
screen "eProC - Seguimiento Datos" 1280x768, template "Template"
   TextField "Campo de texto_9" at 88,77 size 35x18; Text 'Araña'
   TextField "Campo de texto_10" at 265,77 size 32x18; Text 'Rolos'
   TextField "Campo de texto_11" at 439,77 size 54x18; Text 'Perfilador'
   TextField "Campo de texto_12" at 788,77 size 31x18; Text 'Pinza'
   TextField "Campo de texto_13" at 967,77 size 57x18; Text 'Plegadora'
   TextField "Campo de texto_16" at 88,130 size 12x18; Text 'A'
   IOField "Champ E/S_8" at 109,127 size 54x25; FormatPattern 9999999
      Appearance <- "Araña\Araña.PresenciaPieza"
      ProcessValue <- "Araña\Araña.A"
   IOField "Champ E/S_9" at 109,147 size 54x25; FormatPattern 9999999
      Appearance <- "Araña\Araña.PresenciaPieza"
      ProcessValue <- "Araña\Araña.B"
   IOField "Champ E/S_10" at 109,168 size 54x24; FormatPattern 9999999
      Appearance <- "Araña\Araña.PresenciaPieza"
      ProcessValue <- "Araña\Araña.C"
   IOField "Champ E/S_11" at 109,187 size 54x25; FormatPattern 9999999
      Appearance <- "Araña\Araña.PresenciaPieza"
      ProcessValue <- "Araña\Araña.D"
   TextField "Campo de texto_17" at 89,148 size 11x18; Text 'B'
   TextField "Campo de texto_18" at 89,168 size 11x18; Text 'C'
   TextField "Campo de texto_19" at 89,188 size 12x18; Text 'D'
   TextField "Campo de texto_20" at 265,131 size 12x18; Text 'A'
   IOField "Champ E/S_12" at 284,127 size 54x25; FormatPattern 9999999
      Appearance <- "Rolos\Rolos.PresenciaPieza"
      ProcessValue <- "Rolos\Rolos.A"
   IOField "Champ E/S_13" at 284,147 size 54x25; FormatPattern 9999999
      Appearance <- "Rolos\Rolos.PresenciaPieza"
      ProcessValue <- "Rolos\Rolos.B"
   IOField "Champ E/S_14" at 284,168 size 54x24; FormatPattern 9999999
      Appearance <- "Rolos\Rolos.PresenciaPieza"
      ProcessValue <- "Rolos\Rolos.C"
   IOField "Champ E/S_15" at 284,187 size 54x25; FormatPattern 9999999
      Appearance <- "Rolos\Rolos.PresenciaPieza"
      ProcessValue <- "Rolos\Rolos.D"
   TextField "Campo de texto_21" at 265,149 size 11x18; Text 'B'
   TextField "Campo de texto_22" at 265,169 size 11x18; Text 'C'
   TextField "Campo de texto_23" at 265,189 size 12x18; Text 'D'
   TextField "Campo de texto_24" at 439,131 size 12x18; Text 'A'
   IOField "Champ E/S_16" at 462,127 size 53x25; FormatPattern 9999999
      Appearance <- "Perfiladores\Perfilador.PresenciaPieza"
      ProcessValue <- "Perfiladores\Perfilador.A"
   IOField "Champ E/S_17" at 462,147 size 53x25; FormatPattern 9999999
      Appearance <- "Perfiladores\Perfilador.PresenciaPieza"
      ProcessValue <- "Perfiladores\Perfilador.B"
   IOField "Champ E/S_18" at 462,168 size 53x24; FormatPattern 9999999
      Appearance <- "Perfiladores\Perfilador.PresenciaPieza"
      ProcessValue <- "Perfiladores\Perfilador.C"
   IOField "Champ E/S_19" at 462,187 size 53x25; FormatPattern 9999999
      Appearance <- "Perfiladores\Perfilador.PresenciaPieza"
      ProcessValue <- "Perfiladores\Perfilador.D"
   TextField "Campo de texto_25" at 441,149 size 11x18; Text 'B'
   TextField "Campo de texto_26" at 441,169 size 11x18; Text 'C'
   TextField "Campo de texto_27" at 441,189 size 12x18; Text 'D'
   TextField "Campo de texto_28" at 788,131 size 12x18; Text 'A'
   IOField "Champ E/S_20" at 813,127 size 53x25; FormatPattern 9999999
      Appearance <- "Pinza\Pinza.PresenciaPieza"
      ProcessValue <- "Pinza\Pinza.A"
   IOField "Champ E/S_21" at 813,147 size 53x25; FormatPattern 9999999
      Appearance <- "Pinza\Pinza.PresenciaPieza"
      ProcessValue <- "Pinza\Pinza.B"
   IOField "Champ E/S_22" at 813,168 size 53x24; FormatPattern 9999999
      Appearance <- "Pinza\Pinza.PresenciaPieza"
      ProcessValue <- "Pinza\Pinza.C"
   IOField "Champ E/S_23" at 813,187 size 53x25; FormatPattern 9999999
      Appearance <- "Pinza\Pinza.PresenciaPieza"
      ProcessValue <- "Pinza\Pinza.D"
   TextField "Campo de texto_29" at 788,149 size 11x18; Text 'B'
   TextField "Campo de texto_30" at 788,169 size 11x18; Text 'C'
   TextField "Campo de texto_31" at 788,189 size 12x18; Text 'D'
   TextField "Campo de texto_32" at 967,131 size 12x18; Text 'A'
   IOField "Champ E/S_24" at 988,127 size 53x25; FormatPattern 9999999
      Appearance <- "Plegadora\Plegadora.PresenciaPieza"
      ProcessValue <- "Plegadora\Plegadora.A"
   IOField "Champ E/S_25" at 988,147 size 53x25; FormatPattern 9999999
      Appearance <- "Plegadora\Plegadora.PresenciaPieza"
      ProcessValue <- "Plegadora\Plegadora.B"
   IOField "Champ E/S_26" at 988,168 size 53x24; FormatPattern 9999999
      Appearance <- "Plegadora\Plegadora.PresenciaPieza"
      ProcessValue <- "Plegadora\Plegadora.C"
   IOField "Champ E/S_27" at 988,187 size 53x25; FormatPattern 9999999
      Appearance <- "Plegadora\Plegadora.PresenciaPieza"
      ProcessValue <- "Plegadora\Plegadora.D"
   TextField "Campo de texto_33" at 967,149 size 11x18; Text 'B'
   TextField "Campo de texto_34" at 967,169 size 11x18; Text 'C'
   TextField "Campo de texto_35" at 967,189 size 12x18; Text 'D'
   Button "Botón_8" at 437,38 size 80x36; TextOff 'Borrar'; PictureOff "Borrar Pulsador"
      on Click: ResetBit("Perfiladores\Perfilador.PresenciaPieza")
      Visibility <- "Perfiladores\Perfilador.PresenciaPieza"
   Button "Botón_9" at 263,38 size 80x36; TextOff 'Borrar'; PictureOff "Borrar Pulsador"
      on Click: ResetBit("Rolos\Rolos.PresenciaPieza")
      Visibility <- "Rolos\Rolos.PresenciaPieza"
   Button "Botón_10" at 86,38 size 80x36; TextOff 'Borrar'; PictureOff "Borrar Pulsador"
      on Click: ResetBit("Araña\Araña.PresenciaPieza")
      Visibility <- "Araña\Araña.PresenciaPieza"
   TextField "Campo de texto_113" at 615,77 size 31x18; Text 'Cinta'
   TextField "Campo de texto_114" at 615,131 size 12x18; Text 'A'
   IOField "Champ E/S_106" at 638,127 size 53x25; FormatPattern 9999999
      Appearance <- "Cinta\Cinta.PresenciaPieza"
      ProcessValue <- "Cinta\Cinta.A"
   IOField "Champ E/S_107" at 638,147 size 53x25; FormatPattern 9999999
      Appearance <- "Cinta\Cinta.PresenciaPieza"
      ProcessValue <- "Cinta\Cinta.B"
   IOField "Champ E/S_108" at 638,168 size 53x24; FormatPattern 9999999
      Appearance <- "Cinta\Cinta.PresenciaPieza"
      ProcessValue <- "Cinta\Cinta.C"
   IOField "Champ E/S_109" at 638,187 size 53x25; FormatPattern 9999999
      Appearance <- "Cinta\Cinta.PresenciaPieza"
      ProcessValue <- "Cinta\Cinta.D"
   TextField "Campo de texto_115" at 615,149 size 11x18; Text 'B'
   TextField "Campo de texto_116" at 615,169 size 11x18; Text 'C'
   TextField "Campo de texto_117" at 615,189 size 12x18; Text 'D'
   Button "Botón_14" at 613,38 size 80x36; TextOff 'Borrar'; PictureOff "Borrar Pulsador"
      on Click: ResetBit("Cinta\Cinta.PresenciaPieza")
      Visibility <- "Cinta\Cinta.PresenciaPieza"
   Button "Botón_15" at 788,38 size 80x36; TextOff 'Borrar'; PictureOff "Borrar Pulsador"
      on Click: ResetBit("Pinza\Pinza.PresenciaPieza")
      Visibility <- "Pinza\Pinza.PresenciaPieza"
   Button "Botón_16" at 963,38 size 80x36; TextOff 'Borrar'; PictureOff "Borrar Pulsador"
      on Click: ResetBit("Plegadora\Plegadora.PresenciaPieza")
      Visibility <- "Plegadora\Plegadora.PresenciaPieza"
   GraphicView "Visor de gráficos_2" at 211,77 size 29x29; Picture "Gráfico_4"
   GraphicView "Visor de gráficos_1" at 384,77 size 29x29; Picture "Gráfico_4"
   GraphicView "Visor de gráficos_3" at 561,77 size 29x29; Picture "Gráfico_4"
   GraphicView "Visor de gráficos_4" at 734,77 size 29x29; Picture "Gráfico_4"
   GraphicView "Visor de gráficos_5" at 909,77 size 29x29; Picture "Gráfico_4"
   TextField "Campo de texto_1" at 72,425 size 54x29; Text 'Pinza'
   TextField "Campo de texto_2" at 229,507 size 54x18; Text 'Solicitada'
   TextField "Campo de texto_49" at 142,529 size 60x18; Text 'Recepción'
   IOField "Champ E/S_1" at 221,525 size 85x25; FormatPattern s9999999999
      ProcessValue <- "Pos_Recepcion"
      Appearance <- "Pinza\Pinza.PresenciaPieza"
   IOField "Champ E/S_2" at 221,545 size 85x25; FormatPattern s9999999999
      ProcessValue <- "Pos_E1H1"
      Appearance <- "Pinza\Pinza.PresenciaPieza"
   IOField "Champ E/S_3" at 221,566 size 85x24; FormatPattern s9999999999
      ProcessValue <- "Pos_E1H2"
      Appearance <- "Pinza\Pinza.PresenciaPieza"
   IOField "Champ E/S_4" at 221,585 size 85x25; FormatPattern s9999999999
      ProcessValue <- "Pos_E2H1"
      Appearance <- "Pinza\Pinza.PresenciaPieza"
   TextField "Campo de texto_50" at 142,547 size 33x18; Text 'E1H1'
   TextField "Campo de texto_51" at 142,567 size 33x18; Text 'E1H2'
   TextField "Campo de texto_52" at 142,587 size 33x18; Text 'E2H1'
   TextField "Campo de texto_53" at 313,507 size 57x18; Text 'Alcanzada'
   IOField "Champ E/S_5" at 305,525 size 85x25; FormatPattern s9999999999
      ProcessValue <- "Pos_Recepcion(3)"
      Appearance <- "Pinza\Pinza.PresenciaPieza"
   IOField "Champ E/S_6" at 305,545 size 85x25; FormatPattern s9999999999
      ProcessValue <- "Pos_E1H1(3)"
      Appearance <- "Pinza\Pinza.PresenciaPieza"
   IOField "Champ E/S_7" at 305,566 size 85x24; FormatPattern s9999999999
      ProcessValue <- "Pos_E1H2(3)"
      Appearance <- "Pinza\Pinza.PresenciaPieza"
   IOField "Champ E/S_28" at 305,585 size 85x25; FormatPattern s9999999999
      ProcessValue <- "Pos_E2H1(3)"
      Appearance <- "Pinza\Pinza.PresenciaPieza"
   TextField "Campo de texto_65" at 615,507 size 54x18; Text 'Solicitada'
   IOField "Champ E/S_57" at 608,525 size 85x25; FormatPattern s9999999999
      ProcessValue <- "Pos_Recepcion(1)"
      Appearance <- "Pinza\Pinza.PresenciaPieza"
   IOField "Champ E/S_58" at 608,545 size 85x25; FormatPattern s9999999999
      ProcessValue <- "Pos_E1H1(1)"
      Appearance <- "Pinza\Pinza.PresenciaPieza"
   IOField "Champ E/S_59" at 608,566 size 85x24; FormatPattern s9999999999
      ProcessValue <- "Pos_E1H2(1)"
      Appearance <- "Pinza\Pinza.PresenciaPieza"
   IOField "Champ E/S_60" at 608,585 size 85x25; FormatPattern s9999999999
      ProcessValue <- "Pos_E2H1(1)"
      Appearance <- "Pinza\Pinza.PresenciaPieza"
   TextField "Campo de texto_78" at 697,507 size 57x18; Text 'Alcanzada'
   IOField "Champ E/S_69" at 690,525 size 85x25; FormatPattern s9999999999
      ProcessValue <- "Pos_Recepcion(4)"
      Appearance <- "Pinza\Pinza.PresenciaPieza"
   IOField "Champ E/S_70" at 690,545 size 85x25; FormatPattern s9999999999
      ProcessValue <- "Pos_E1H1(4)"
      Appearance <- "Pinza\Pinza.PresenciaPieza"
   IOField "Champ E/S_71" at 690,566 size 85x24; FormatPattern s9999999999
      ProcessValue <- "Pos_E1H2(4)"
      Appearance <- "Pinza\Pinza.PresenciaPieza"
   IOField "Champ E/S_72" at 690,585 size 85x25; FormatPattern s9999999999
      ProcessValue <- "Pos_E2H1(4)"
      Appearance <- "Pinza\Pinza.PresenciaPieza"
   TextField "Campo de texto_91" at 1003,507 size 54x18; Text 'Solicitada'
   IOField "Champ E/S_81" at 995,525 size 85x25; FormatPattern s9999999999
      ProcessValue <- "Pos_Recepcion(2)"
      Appearance <- "Pinza\Pinza.PresenciaPieza"
   IOField "Champ E/S_82" at 995,545 size 85x25; FormatPattern s9999999999
      ProcessValue <- "Pos_E1H1(2)"
      Appearance <- "Pinza\Pinza.PresenciaPieza"
   IOField "Champ E/S_83" at 995,566 size 85x24; FormatPattern s9999999999
      ProcessValue <- "Pos_E1H2(2)"
      Appearance <- "Pinza\Pinza.PresenciaPieza"
   IOField "Champ E/S_84" at 995,585 size 85x25; FormatPattern s9999999999
      ProcessValue <- "Pos_E2H1(2)"
      Appearance <- "Pinza\Pinza.PresenciaPieza"
   TextField "Campo de texto_104" at 1085,507 size 57x18; Text 'Alcanzada'
   IOField "Champ E/S_93" at 1077,525 size 85x25; FormatPattern s9999999999
      ProcessValue <- "Pos_Recepcion(5)"
      Appearance <- "Pinza\Pinza.PresenciaPieza"
   IOField "Champ E/S_94" at 1077,545 size 85x25; FormatPattern s9999999999
      ProcessValue <- "Pos_E1H1(5)"
      Appearance <- "Pinza\Pinza.PresenciaPieza"
   IOField "Champ E/S_95" at 1077,566 size 85x24; FormatPattern s9999999999
      ProcessValue <- "Pos_E1H2(5)"
      Appearance <- "Pinza\Pinza.PresenciaPieza"
   IOField "Champ E/S_96" at 1077,585 size 85x25; FormatPattern s9999999999
      ProcessValue <- "Pos_E2H1(5)"
      Appearance <- "Pinza\Pinza.PresenciaPieza"
   TextField "Campo de texto_55" at 533,529 size 60x18; Text 'Recepción'
   TextField "Campo de texto_56" at 533,547 size 33x18; Text 'E1H1'
   TextField "Campo de texto_57" at 533,567 size 33x18; Text 'E1H2'
   TextField "Campo de texto_58" at 533,587 size 33x18; Text 'E2H1'
   TextField "Campo de texto_59" at 916,529 size 60x18; Text 'Recepción'
   TextField "Campo de texto_60" at 916,547 size 33x18; Text 'E1H1'
   TextField "Campo de texto_61" at 916,567 size 33x18; Text 'E1H2'
   TextField "Campo de texto_62" at 916,587 size 33x18; Text 'E2H1'
   TextField "Campo de texto_63" at 231,488 size 128x18; Text 'Posición pieza anterior:'
   TextField "Campo de texto_64" at 616,488 size 139x18; Text 'Posición pieza anterior 2:'
   TextField "Campo de texto_66" at 1002,488 size 139x18; Text 'Posición pieza anterior 3:'
   Button "Template_Plantilla_Botón_33" at 275,715 size 150x53; TextOff 'SEGUIMIENTO DE DATOS'
   Button "Template_Plantilla_Bouton_2" at 1085,715 size 193x53; TextOff 'ALARMAS / DEFAUT'
      on Press: ActivateScreen("eProC - Alarmas", 0)
      Visibility <- "DB_OP.P_DEFAUT"
   TextField "Campo de texto_3" at 1138,77 size 71x18; Text 'Descargador'
   TextField "Campo de texto_4" at 1138,131 size 13x18; Text 'A'
   IOField "Champ E/S_37" at 1159,127 size 54x25; FormatPattern 9999999
      ProcessValue <- "Descargador-A"
      Appearance <- "Descargador-PiezaPresente"
   IOField "Champ E/S_38" at 1159,147 size 54x25; FormatPattern 9999999
      ProcessValue <- "Descargador-B"
      Appearance <- "Descargador-PiezaPresente"
   IOField "Champ E/S_39" at 1159,168 size 54x24; FormatPattern 9999999
      ProcessValue <- "Descargador-C"
      Appearance <- "Descargador-PiezaPresente"
   IOField "Champ E/S_40" at 1159,187 size 54x25; FormatPattern 9999999
      ProcessValue <- "Descargador-D"
      Appearance <- "Descargador-PiezaPresente"
   TextField "Campo de texto_5" at 1138,149 size 12x18; Text 'B'
   TextField "Campo de texto_6" at 1138,169 size 12x18; Text 'C'
   TextField "Campo de texto_7" at 1138,189 size 13x18; Text 'D'
   Button "Botón_1" at 1134,38 size 81x36; TextOff 'Borrar'; PictureOff "Borrar Pulsador"
      on Click: ResetBit("Descargador-PiezaPresente")
      Visibility <- "Descargador-PiezaPresente"
   GraphicView "Visor de gráficos_6" at 1080,77 size 30x29; Picture "Gráfico_4"
   TextField "Campo de texto_118" at 441,210 size 17x18; Text 'F1'
   IOField "Champ E/S_110" at 465,207 size 51x25; FormatPattern s999999
      Appearance <- "Perfiladores\Perfilador.PresenciaPieza"
      ProcessValue <- "Perfiladores\Perfilador.F1"
   IOField "Champ E/S_111" at 465,227 size 51x25; FormatPattern s999999
      Appearance <- "Perfiladores\Perfilador.PresenciaPieza"
      ProcessValue <- "Perfiladores\Perfilador.F2"
   IOField "Champ E/S_112" at 465,248 size 51x24; FormatPattern s999999
      Appearance <- "Perfiladores\Perfilador.PresenciaPieza"
      ProcessValue <- "Perfiladores\Perfilador.F3"
   IOField "Champ E/S_113" at 465,267 size 51x25; FormatPattern s999999
      Appearance <- "Perfiladores\Perfilador.PresenciaPieza"
      ProcessValue <- "Perfiladores\Perfilador.F4"
   TextField "Campo de texto_119" at 441,229 size 17x18; Text 'F2'
   TextField "Campo de texto_120" at 441,249 size 17x18; Text 'F3'
   TextField "Campo de texto_121" at 441,269 size 17x18; Text 'F4'
   TextField "Campo de texto_122" at 441,290 size 35x18; Text 'PL1-1'
   IOField "Champ E/S_114" at 481,287 size 51x25; FormatPattern s999999
      Appearance <- "Perfiladores\Perfilador.PresenciaPieza"
      ProcessValue <- "Perfiladores\Perfilador.PL1_1"
   IOField "Champ E/S_115" at 481,307 size 51x25; FormatPattern s999999
      Appearance <- "Perfiladores\Perfilador.PresenciaPieza"
      ProcessValue <- "Perfiladores\Perfilador.PL1_2"
   IOField "Champ E/S_116" at 481,328 size 51x24; FormatPattern s999999
      Appearance <- "Perfiladores\Perfilador.PresenciaPieza"
      ProcessValue <- "Perfiladores\Perfilador.PL2_1"
   IOField "Champ E/S_117" at 481,347 size 51x25; FormatPattern s999999
      Appearance <- "Perfiladores\Perfilador.PresenciaPieza"
      ProcessValue <- "Perfiladores\Perfilador.PL2_2"
   TextField "Campo de texto_123" at 441,310 size 35x18; Text 'PL1-2'
   TextField "Campo de texto_124" at 441,331 size 35x18; Text 'PL2-1'
   TextField "Campo de texto_125" at 441,350 size 35x18; Text 'PL2-2'
   TextField "Campo de texto_134" at 266,210 size 17x18; Text 'F1'
   IOField "Champ E/S_126" at 290,207 size 51x25; FormatPattern s999999
      Appearance <- "Rolos\Rolos.PresenciaPieza"
      ProcessValue <- "Rolos\Rolos.F1"
   IOField "Champ E/S_127" at 290,227 size 51x25; FormatPattern s999999
      Appearance <- "Rolos\Rolos.PresenciaPieza"
      ProcessValue <- "Rolos\Rolos.F2"
   IOField "Champ E/S_128" at 290,248 size 51x24; FormatPattern s999999
      Appearance <- "Rolos\Rolos.PresenciaPieza"
      ProcessValue <- "Rolos\Rolos.F3"
   IOField "Champ E/S_129" at 290,267 size 51x25; FormatPattern s999999
      Appearance <- "Rolos\Rolos.PresenciaPieza"
      ProcessValue <- "Rolos\Rolos.F4"
   TextField "Campo de texto_135" at 266,229 size 17x18; Text 'F2'
   TextField "Campo de texto_136" at 266,249 size 17x18; Text 'F3'
   TextField "Campo de texto_137" at 266,269 size 17x18; Text 'F4'
   TextField "Campo de texto_138" at 266,290 size 35x18; Text 'PL1-1'
   IOField "Champ E/S_130" at 306,287 size 51x25; FormatPattern s999999
      Appearance <- "Rolos\Rolos.PresenciaPieza"
      ProcessValue <- "Rolos\Rolos.PL1_1"
   IOField "Champ E/S_131" at 306,307 size 51x25; FormatPattern s999999
      Appearance <- "Rolos\Rolos.PresenciaPieza"
      ProcessValue <- "Rolos\Rolos.PL1_2"
   IOField "Champ E/S_132" at 306,328 size 51x24; FormatPattern s999999
      Appearance <- "Rolos\Rolos.PresenciaPieza"
      ProcessValue <- "Rolos\Rolos.PL2_1"
   IOField "Champ E/S_133" at 306,347 size 51x25; FormatPattern s999999
      Appearance <- "Rolos\Rolos.PresenciaPieza"
      ProcessValue <- "Rolos\Rolos.PL2_2"
   TextField "Campo de texto_139" at 266,310 size 35x18; Text 'PL1-2'
   TextField "Campo de texto_140" at 266,331 size 35x18; Text 'PL2-1'
   TextField "Campo de texto_141" at 266,350 size 35x18; Text 'PL2-2'
   TextField "Campo de texto_142" at 89,210 size 17x18; Text 'F1'
   IOField "Champ E/S_134" at 113,207 size 51x25; FormatPattern s999999
      Appearance <- "Araña\Araña.PresenciaPieza"
      ProcessValue <- "Araña\Araña.F1"
   IOField "Champ E/S_135" at 113,227 size 51x25; FormatPattern s999999
      Appearance <- "Araña\Araña.PresenciaPieza"
      ProcessValue <- "Araña\Araña.F2"
   IOField "Champ E/S_136" at 113,248 size 51x24; FormatPattern s999999
      Appearance <- "Araña\Araña.PresenciaPieza"
      ProcessValue <- "Araña\Araña.F3"
   IOField "Champ E/S_137" at 113,267 size 51x25; FormatPattern s999999
      Appearance <- "Araña\Araña.PresenciaPieza"
      ProcessValue <- "Araña\Araña.F4"
   TextField "Campo de texto_143" at 89,229 size 17x18; Text 'F2'
   TextField "Campo de texto_144" at 89,249 size 17x18; Text 'F3'
   TextField "Campo de texto_145" at 89,269 size 17x18; Text 'F4'
   TextField "Campo de texto_146" at 89,290 size 35x18; Text 'PL1-1'
   IOField "Champ E/S_138" at 129,287 size 51x25; FormatPattern s999999
      Appearance <- "Araña\Araña.PresenciaPieza"
      ProcessValue <- "Araña\Araña.PL1_1"
   IOField "Champ E/S_139" at 129,307 size 51x25; FormatPattern s999999
      Appearance <- "Araña\Araña.PresenciaPieza"
      ProcessValue <- "Araña\Araña.PL1_2"
   IOField "Champ E/S_140" at 129,328 size 51x24; FormatPattern s999999
      Appearance <- "Araña\Araña.PresenciaPieza"
      ProcessValue <- "Araña\Araña.PL2_1"
   IOField "Champ E/S_141" at 129,347 size 51x25; FormatPattern s999999
      Appearance <- "Araña\Araña.PresenciaPieza"
      ProcessValue <- "Araña\Araña.PL2_2"
   TextField "Campo de texto_147" at 89,310 size 35x18; Text 'PL1-2'
   TextField "Campo de texto_148" at 89,331 size 35x18; Text 'PL2-1'
   TextField "Campo de texto_149" at 89,350 size 35x18; Text 'PL2-2'
   TextField "Campo de texto_150" at 617,210 size 17x18; Text 'F1'
   IOField "Champ E/S_142" at 641,207 size 51x25; FormatPattern s999999
      Appearance <- "Cinta\Cinta.PresenciaPieza"
      ProcessValue <- "Cinta\Cinta.F1"
   IOField "Champ E/S_143" at 641,227 size 51x25; FormatPattern s999999
      Appearance <- "Cinta\Cinta.PresenciaPieza"
      ProcessValue <- "Cinta\Cinta.F2"
   IOField "Champ E/S_144" at 641,248 size 51x24; FormatPattern s999999
      Appearance <- "Cinta\Cinta.PresenciaPieza"
      ProcessValue <- "Cinta\Cinta.F3"
   IOField "Champ E/S_145" at 641,267 size 51x25; FormatPattern s999999
      Appearance <- "Cinta\Cinta.PresenciaPieza"
      ProcessValue <- "Cinta\Cinta.F4"
   TextField "Campo de texto_151" at 617,229 size 17x18; Text 'F2'
   TextField "Campo de texto_152" at 617,249 size 17x18; Text 'F3'
   TextField "Campo de texto_153" at 617,269 size 17x18; Text 'F4'
   TextField "Campo de texto_154" at 617,290 size 35x18; Text 'PL1-1'
   IOField "Champ E/S_146" at 657,287 size 51x25; FormatPattern s999999
      Appearance <- "Cinta\Cinta.PresenciaPieza"
      ProcessValue <- "Cinta\Cinta.PL1_1"
   IOField "Champ E/S_147" at 657,307 size 51x25; FormatPattern s999999
      Appearance <- "Cinta\Cinta.PresenciaPieza"
      ProcessValue <- "Cinta\Cinta.PL1_2"
   IOField "Champ E/S_148" at 657,328 size 51x24; FormatPattern s999999
      Appearance <- "Cinta\Cinta.PresenciaPieza"
      ProcessValue <- "Cinta\Cinta.PL2_1"
   IOField "Champ E/S_149" at 657,347 size 51x25; FormatPattern s999999
      Appearance <- "Cinta\Cinta.PresenciaPieza"
      ProcessValue <- "Cinta\Cinta.PL2_2"
   TextField "Campo de texto_155" at 617,310 size 35x18; Text 'PL1-2'
   TextField "Campo de texto_156" at 617,331 size 35x18; Text 'PL2-1'
   TextField "Campo de texto_157" at 617,350 size 35x18; Text 'PL2-2'
   TextField "Campo de texto_158" at 789,210 size 17x18; Text 'F1'
   IOField "Champ E/S_150" at 813,207 size 51x25; FormatPattern s999999
      Appearance <- "Pinza\Pinza.PresenciaPieza"
      ProcessValue <- "Pinza\Pinza.F1"
   IOField "Champ E/S_151" at 813,227 size 51x25; FormatPattern s999999
      Appearance <- "Pinza\Pinza.PresenciaPieza"
      ProcessValue <- "Pinza\Pinza.F2"
   IOField "Champ E/S_152" at 813,248 size 51x24; FormatPattern s999999
      Appearance <- "Pinza\Pinza.PresenciaPieza"
      ProcessValue <- "Pinza\Pinza.F3"
   IOField "Champ E/S_153" at 813,267 size 51x25; FormatPattern s999999
      Appearance <- "Pinza\Pinza.PresenciaPieza"
      ProcessValue <- "Pinza\Pinza.F4"
   TextField "Campo de texto_159" at 789,229 size 17x18; Text 'F2'
   TextField "Campo de texto_160" at 789,249 size 17x18; Text 'F3'
   TextField "Campo de texto_161" at 789,269 size 17x18; Text 'F4'
   TextField "Campo de texto_162" at 789,290 size 35x18; Text 'PL1-1'
   IOField "Champ E/S_154" at 829,287 size 51x25; FormatPattern s999999
      Appearance <- "Pinza\Pinza.PresenciaPieza"
      ProcessValue <- "Pinza\Pinza.PL1_1"
   IOField "Champ E/S_155" at 829,307 size 51x25; FormatPattern s999999
      Appearance <- "Pinza\Pinza.PresenciaPieza"
      ProcessValue <- "Pinza\Pinza.PL1_2"
   IOField "Champ E/S_156" at 829,328 size 51x24; FormatPattern s999999
      Appearance <- "Pinza\Pinza.PresenciaPieza"
      ProcessValue <- "Pinza\Pinza.PL2_1"
   IOField "Champ E/S_157" at 829,347 size 51x25; FormatPattern s999999
      Appearance <- "Pinza\Pinza.PresenciaPieza"
      ProcessValue <- "Pinza\Pinza.PL2_2"
   TextField "Campo de texto_163" at 789,310 size 35x18; Text 'PL1-2'
   TextField "Campo de texto_164" at 789,331 size 35x18; Text 'PL2-1'
   TextField "Campo de texto_165" at 789,350 size 35x18; Text 'PL2-2'
   TextField "Campo de texto_166" at 967,210 size 17x18; Text 'F1'
   IOField "Champ E/S_158" at 991,207 size 51x25; FormatPattern s999999
      Appearance <- "Plegadora\Plegadora.PresenciaPieza"
      ProcessValue <- "Plegadora\Plegadora.F1"
   IOField "Champ E/S_159" at 991,227 size 51x25; FormatPattern s999999
      Appearance <- "Plegadora\Plegadora.PresenciaPieza"
      ProcessValue <- "Plegadora\Plegadora.F2"
   IOField "Champ E/S_160" at 991,248 size 51x24; FormatPattern s999999
      Appearance <- "Plegadora\Plegadora.PresenciaPieza"
      ProcessValue <- "Plegadora\Plegadora.F3"
   IOField "Champ E/S_161" at 991,267 size 51x25; FormatPattern s999999
      Appearance <- "Plegadora\Plegadora.PresenciaPieza"
      ProcessValue <- "Plegadora\Plegadora.F4"
   TextField "Campo de texto_167" at 967,229 size 17x18; Text 'F2'
   TextField "Campo de texto_168" at 967,249 size 17x18; Text 'F3'
   TextField "Campo de texto_169" at 967,269 size 17x18; Text 'F4'
   TextField "Campo de texto_170" at 967,290 size 35x18; Text 'PL1-1'
   IOField "Champ E/S_162" at 1007,287 size 51x25; FormatPattern s999999
      Appearance <- "Plegadora\Plegadora.PresenciaPieza"
      ProcessValue <- "Plegadora\Plegadora.PL1_1"
   IOField "Champ E/S_163" at 1007,307 size 51x25; FormatPattern s999999
      Appearance <- "Plegadora\Plegadora.PresenciaPieza"
      ProcessValue <- "Plegadora\Plegadora.PL1_2"
   IOField "Champ E/S_164" at 1007,328 size 51x24; FormatPattern s999999
      Appearance <- "Plegadora\Plegadora.PresenciaPieza"
      ProcessValue <- "Plegadora\Plegadora.PL2_1"
   IOField "Champ E/S_165" at 1007,347 size 51x25; FormatPattern s999999
      Appearance <- "Plegadora\Plegadora.PresenciaPieza"
      ProcessValue <- "Plegadora\Plegadora.PL2_2"
   TextField "Campo de texto_171" at 967,310 size 35x18; Text 'PL1-2'
   TextField "Campo de texto_172" at 967,331 size 35x18; Text 'PL2-1'
   TextField "Campo de texto_173" at 967,350 size 35x18; Text 'PL2-2'
   IOField "Champ E/S_32" at 443,100 size 80x25; FormatPattern ????????????????????
      Appearance <- "Perfiladores\Perfilador.PresenciaPieza"
      ProcessValue <- "Perfiladores\Perfilador.Nombre"
   IOField "Champ E/S_33" at 268,100 size 80x25; FormatPattern ????????????????????
      Appearance <- "Rolos\Rolos.PresenciaPieza"
      ProcessValue <- "Rolos\Rolos.Nombre"
   IOField "Champ E/S_34" at 91,100 size 80x25; FormatPattern ????????????????????
      Appearance <- "Araña\Araña.PresenciaPieza"
      ProcessValue <- "Araña\Araña.Nombre"
   IOField "Champ E/S_35" at 619,100 size 80x25; FormatPattern ????????????????????
      Appearance <- "Cinta\Cinta.PresenciaPieza"
      ProcessValue <- "Cinta\Cinta.Nombre"
   IOField "Champ E/S_41" at 791,100 size 80x25; FormatPattern ????????????????????
      Appearance <- "Pinza\Pinza.PresenciaPieza"
      ProcessValue <- "Pinza\Pinza.Nombre"
   IOField "Champ E/S_42" at 969,100 size 80x25; FormatPattern ????????????????????
      Appearance <- "Plegadora\Plegadora.PresenciaPieza"
      ProcessValue <- "Plegadora\Plegadora.Nombre"
   TextField "Campo de texto_67" at 143,608 size 33x18; Text 'E2H2'
   IOField "Champ E/S_29" at 221,605 size 85x25; FormatPattern s9999999999
      ProcessValue <- "Pos_E2H2"
      Appearance <- "Pinza\Pinza.PresenciaPieza"
   IOField "Champ E/S_30" at 221,625 size 85x25; FormatPattern s9999999999
      ProcessValue <- "Pos_Entrega"
      Appearance <- "Pinza\Pinza.PresenciaPieza"
   TextField "Campo de texto_68" at 143,627 size 47x18; Text 'Entrega'
   IOField "Champ E/S_31" at 305,605 size 85x25; FormatPattern s9999999999
      ProcessValue <- "Pos_E2H2(3)"
      Appearance <- "Pinza\Pinza.PresenciaPieza"
   IOField "Champ E/S_36" at 305,625 size 85x25; FormatPattern s9999999999
      ProcessValue <- "Pos_Entrega(3)"
      Appearance <- "Pinza\Pinza.PresenciaPieza"
   IOField "Champ E/S_61" at 608,605 size 85x25; FormatPattern s9999999999
      ProcessValue <- "Pos_E2H2(1)"
      Appearance <- "Pinza\Pinza.PresenciaPieza"
   IOField "Champ E/S_62" at 608,625 size 85x25; FormatPattern s9999999999
      ProcessValue <- "Pos_Entrega(1)"
      Appearance <- "Pinza\Pinza.PresenciaPieza"
   IOField "Champ E/S_73" at 690,605 size 85x25; FormatPattern s9999999999
      ProcessValue <- "Pos_E2H2(4)"
      Appearance <- "Pinza\Pinza.PresenciaPieza"
   IOField "Champ E/S_74" at 690,625 size 85x25; FormatPattern s9999999999
      ProcessValue <- "Pos_Entrega(4)"
      Appearance <- "Pinza\Pinza.PresenciaPieza"
   IOField "Champ E/S_85" at 995,605 size 85x25; FormatPattern s9999999999
      ProcessValue <- "Pos_E2H2(2)"
      Appearance <- "Pinza\Pinza.PresenciaPieza"
   IOField "Champ E/S_86" at 995,625 size 85x25; FormatPattern s9999999999
      ProcessValue <- "Pos_Entrega(2)"
      Appearance <- "Pinza\Pinza.PresenciaPieza"
   IOField "Champ E/S_97" at 1077,605 size 85x25; FormatPattern s9999999999
      ProcessValue <- "Pos_E2H2(5)"
      Appearance <- "Pinza\Pinza.PresenciaPieza"
   IOField "Champ E/S_98" at 1077,625 size 85x25; FormatPattern s9999999999
      ProcessValue <- "Pos_Entrega(5)"
      Appearance <- "Pinza\Pinza.PresenciaPieza"
   TextField "Campo de texto_69" at 534,608 size 33x18; Text 'E2H2'
   TextField "Campo de texto_70" at 534,627 size 47x18; Text 'Entrega'
   TextField "Campo de texto_71" at 917,608 size 33x18; Text 'E2H2'
   TextField "Campo de texto_72" at 917,627 size 47x18; Text 'Entrega'
   TextField "Campo de texto_8" at 1138,210 size 18x18; Text 'F1'
   IOField "Champ E/S_43" at 1162,207 size 52x25; FormatPattern s999999
      ProcessValue <- "Descargador-F1"
      Appearance <- "Descargador-PiezaPresente"
   IOField "Champ E/S_44" at 1162,227 size 52x25; FormatPattern s999999
      ProcessValue <- "Descargador-F2"
      Appearance <- "Descargador-PiezaPresente"
   IOField "Champ E/S_45" at 1162,248 size 52x24; FormatPattern s999999
      ProcessValue <- "Descargador-F3"
      Appearance <- "Descargador-PiezaPresente"
   IOField "Champ E/S_46" at 1162,267 size 52x25; FormatPattern s999999
      ProcessValue <- "Descargador-F4"
      Appearance <- "Descargador-PiezaPresente"
   TextField "Campo de texto_14" at 1138,229 size 18x18; Text 'F2'
   TextField "Campo de texto_15" at 1138,249 size 18x18; Text 'F3'
   TextField "Campo de texto_36" at 1138,269 size 18x18; Text 'F4'
   TextField "Campo de texto_37" at 1138,290 size 36x18; Text 'PL1-1'
   IOField "Champ E/S_47" at 1178,287 size 52x25; FormatPattern s999999
      ProcessValue <- "Descargador-PL1_1"
      Appearance <- "Descargador-PiezaPresente"
   IOField "Champ E/S_48" at 1178,307 size 52x25; FormatPattern s999999
      ProcessValue <- "Descargador-PL1_2"
      Appearance <- "Descargador-PiezaPresente"
   IOField "Champ E/S_49" at 1178,328 size 52x24; FormatPattern s999999
      ProcessValue <- "Descargador-PL2_1"
      Appearance <- "Descargador-PiezaPresente"
   IOField "Champ E/S_50" at 1178,347 size 52x25; FormatPattern s999999
      ProcessValue <- "Descargador-PL2_2"
      Appearance <- "Descargador-PiezaPresente"
   TextField "Campo de texto_38" at 1138,310 size 36x18; Text 'PL1-2'
   TextField "Campo de texto_39" at 1138,331 size 36x18; Text 'PL2-1'
   TextField "Campo de texto_40" at 1138,350 size 36x18; Text 'PL2-2'
   IOField "Champ E/S_51" at 1140,100 size 81x25; FormatPattern ????????????????????
      ProcessValue <- "Descargador-Nombre"
      Appearance <- "Descargador-PiezaPresente"

Template "Template" 1280x768
   TextField "Template_Plantilla_Campo de texto" at 0,0 size 1280x24; Text 'Movimiento Manual Seleccionado -'
      Visibility <- "DB_OP.RC1"
   TextField "Template_Plantilla_Campo de texto_0" at 0,-1 size 1280x24; Text 'Movimiento Manual Seleccionado -'
      Visibility <- "DB_OP.RC2"
   Button "Template_Plantilla_Bouton_1" at 278,715 size 150x53; TextOff 'SEGUIMIENTO DE DATOS SYSTEM'
      on Click: ActivateScreen("eProC - Seguimiento Datos", 0)
   Button "Template_Plantilla_Bouton_0" at 1085,715 size 193x53; TextOff 'ALARMAS / DEFAUT'
      on Press: ActivateScreen("eProC - Alarmas", 0)
   Button "Template_Plantilla_Botón_2" at 573,715 size 70x53; TextOff 'Text'; Authorization "Nivel 2"; PictureOn "Usuario"; PictureOff "Usuario"
      on Activate: ActivateScreen("Gesión de Usuarios", 0)
   Button "Template_Plantilla_Botón_3" at 129,715 size 150x53; TextOff 'SELECCIÓN RECETAS'
      on Click: ActivateScreen("eProC - Recetas", 0)
   Button "Template_Plantilla_Botón_4" at 641,715 size 150x53; TextOff 'Text'
   SymbolicIOField "Template_Plantilla_Campo ES simbólico" at 234,0 size 896x24; TextOff '0'; TextOn '1'; TextList "RC2"
      ProcessValue <- "DB_OP.RC2"
      Visibility <- "DB_OP.RC2"
   SymbolicIOField "Template_Plantilla_Campo ES simbólico_0" at 234,0 size 896x24; TextOff '0'; TextOn '1'; TextList "RC1"
      ProcessValue <- "DB_OP.RC1"
      Visibility <- "DB_OP.RC1"
   Button "Plantilla_Botón_1" at 1,715 size 130x53; TextOff 'PRINCIPAL'
      on Click: ActivateScreen("eProC - Principal", 0)
   SymbolicIOField "Template_Plantilla_Campo ES simbólico_1" at 0,0 size 1280x24; TextOff '0'; TextOn '1'; TextList "Warnings"
      ProcessValue <- "Warnings"
      Visibility <- "Warning Activo"
   Button "Template_Plantilla_Botón_5" at 789,715 size 150x53; TextOff 'ACUSAR DEFECTO'
      on Click: ActivateScreen("eProC - Defectos", 0)
   Button "Template_Plantilla_Botón_6" at 937,715 size 150x53; TextOff 'Text'
   Button "Template_Plantilla_Bouton_2" at 1085,715 size 193x53; TextOff 'ALARMAS / DEFAUT'
      on Press: ActivateScreen("eProC - Alarmas", 0)
      Visibility <- "DB_OP.P_DEFAUT"
   Button "Template_Plantilla_Botón_1" at 424,715 size 150x53; TextOff 'Text'

PopupScreen "Comandos Araña" 1280x714
   Circle "Cercle_11" at 358,354 size 13x13
      Appearance <- "25S8"
   Circle "Cercle_12" at 359,303 size 13x13
      Appearance <- "25S7"
   Circle "Cercle_0" at 358,375 size 13x13
      Appearance <- "25S4"
   Circle "Cercle_1" at 398,262 size 12x12
      Appearance <- "25S3"
   Circle "Cercle_2" at 320,381 size 12x12
      Appearance <- "25S5"
   Circle "Cercle_3" at 399,300 size 12x12
      Appearance <- "26S3"
   TextField "Campo de texto_1" at 509,184 size 154x18; Text '25S3 - Fin de Carrera Arriba'
   TextField "Campo de texto_6" at 94,362 size 154x18; Text '25S5 - Fin de Carrera Abajo'
   TextField "Campo de texto_10" at 515,231 size 176x18; Text '26S3 - En Posición de Descarga'
   TextField "Campo de texto_8" at 105,226 size 148x18; Text '25S7 - Pistón 2 Expandido'
   TextField "Campo de texto_18" at 107,270 size 144x18; Text '25S8 - Pistón 2 Contraído'
   TextField "Campo de texto_19" at 107,326 size 144x18; Text '25S4 - Pistón 1 Contraído'
   TextField "Campo de texto_20" at 521,268 size 110x18; Text '25S6 - Araña Abajo'
   Circle "Cercle_5" at 401,347 size 13x13
      Appearance <- "25S6"
   Circle "Cercle" at 340,467 size 13x13
      Appearance <- "26S1"
   TextField "Campo de texto_9" at 91,496 size 204x18; Text '26S1 - Tulipas Apoyadas en la Chapa'
   TextField "Campo de texto_21" at 657,356 size 126x18; Text '26S5 - Bajar Velocidad'
   TextField "Campo de texto_22" at 652,316 size 176x18; Text '26S3 - En Posición de Descarga'
   TextField "Campo de texto_23" at 653,421 size 170x46; Text 'M03 - Motor Transporte Araña KM02.1 -> Hacia Rolos KM02.2 -> Hacia Almacenes'
   TextField "Campo de texto_24" at 672,505 size 126x18; Text '26S4 - Bajar Velocidad'
   TextField "Campo de texto_25" at 678,546 size 157x18; Text '26S2 - En Posición de Carga'
   Circle "Cercle_4" at 572,534 size 12x12
      Appearance <- "26S2"
   Circle "Cercle_6" at 567,494 size 12x12
      Appearance <- "26S4"
   Circle "Cercle_7" at 554,342 size 12x12
      Appearance <- "26S5"
   Circle "Cercle_8" at 549,303 size 12x12
      Appearance <- "26S3"
   Polygon "Polígono_3" at 206,439 size 325x50
      Visibility <- "Araña\Araña.PresenciaPieza"
   Rectangle "Rectángulo_7" at 989,250 size 248x208
      Visibility <- "MANU"
   Rectangle "Rectángulo_12" at 989,246 size 248x29
      Visibility <- "MANU"
   Rectangle "Rectángulo_9" at 843,27 size 118x128
      Visibility <- "MANU"
   Rectangle "Rectángulo_8" at 843,27 size 118x29
      Visibility <- "MANU"
   TextField "Campo de texto_3" at 870,31 size 64x18; Text 'Transporte'
      Visibility <- "MANU"
   TextField "Campo de texto_11" at 1010,252 size 66x18; Text 'Aire Tulipas'
      Visibility <- "MANU"
   Button "Botón_4" at 859,71 size 88x33; TextOff 'Avance'
      on Press: SetTag("DB_OP.RC1", 11); SetBit("DB_OP.OP_SELMANU1")
      Visibility <- "MANU"
      Appearance <- "DB_OP.RC1"
   Button "Botón_5" at 859,109 size 88x33; TextOff 'Retroceso'
      on Press: SetTag("DB_OP.RC1", 12); SetBit("DB_OP.OP_SELMANU1")
      Visibility <- "MANU"
      Appearance <- "DB_OP.RC1"
   Button "Botón_10" at 1065,290 size 72x33; TextOff 'Activar'
      on Press: SetTag("DB_OP.RC1", 20); SetBit("DB_OP.OP_SELMANU1")
      Visibility <- "MANU"
      Appearance <- "DB_OP.RC1"
   Button "Botón_17" at 1145,290 size 72x33; TextOff 'Desactivar'
      on Press: SetTag("DB_OP.RC1", 21); SetBit("DB_OP.OP_SELMANU1")
      Visibility <- "MANU"
      Appearance <- "DB_OP.RC1"
   TextField "Campo de texto_12" at 1010,296 size 37x18; Text 'Todas'
      Visibility <- "MANU"
   Button "Botón_1" at 1065,336 size 72x33; TextOff 'Activar'
      on Press: SetTag("DB_OP.RC1", 32); SetBit("DB_OP.OP_SELMANU1")
      Visibility <- "MANU"
      Appearance <- "DB_OP.RC1"
   Button "Botón_23" at 1065,373 size 72x33; TextOff 'Activar'
      on Press: SetTag("DB_OP.RC1", 34); SetBit("DB_OP.OP_SELMANU1")
      Visibility <- "MANU"
      Appearance <- "DB_OP.RC1"
   Button "Botón_24" at 1065,411 size 72x33; TextOff 'Activar'
      on Press: SetTag("DB_OP.RC1", 36); SetBit("DB_OP.OP_SELMANU1")
      Visibility <- "MANU"
      Appearance <- "DB_OP.RC1"
   Button "Botón_26" at 1145,336 size 72x33; TextOff 'Desactivar'
      on Press: SetTag("DB_OP.RC1", 33); SetBit("DB_OP.OP_SELMANU1")
      Visibility <- "MANU"
      Appearance <- "DB_OP.RC1"
   Button "Botón_27" at 1145,373 size 72x33; TextOff 'Desactivar'
      on Press: SetTag("DB_OP.RC1", 35); SetBit("DB_OP.OP_SELMANU1")
      Visibility <- "MANU"
      Appearance <- "DB_OP.RC1"
   Button "Botón_28" at 1145,411 size 72x33; TextOff 'Desactivar'
      on Press: SetTag("DB_OP.RC1", 37); SetBit("DB_OP.OP_SELMANU1")
      Visibility <- "MANU"
      Appearance <- "DB_OP.RC1"
   TextField "Campo de texto_2" at 1008,343 size 48x18; Text 'Grupo 1'
      Visibility <- "MANU"
   TextField "Campo de texto_4" at 1008,381 size 48x18; Text 'Grupo 2'
      Visibility <- "MANU"
   TextField "Campo de texto_5" at 1008,419 size 48x18; Text 'Grupo 3'
      Visibility <- "MANU"
   Rectangle "Rectángulo_1" at 989,483 size 248x208
      Visibility <- "MANU"
   Rectangle "Rectángulo_2" at 989,479 size 248x29
      Visibility <- "MANU"
   TextField "Campo de texto_13" at 1010,485 size 74x18; Text 'Vacío Tulipas'
      Visibility <- "MANU"
   TextField "Campo de texto_14" at 1010,529 size 37x18; Text 'Todas'
      Visibility <- "MANU"
   TextField "Campo de texto_15" at 1008,576 size 48x18; Text 'Grupo 1'
      Visibility <- "MANU"
   TextField "Campo de texto_16" at 1008,614 size 48x18; Text 'Grupo 2'
      Visibility <- "MANU"
   TextField "Campo de texto_17" at 1008,652 size 48x18; Text 'Grupo 3'
      Visibility <- "MANU"
   Button "Botón_21" at 1065,523 size 72x33; TextOff 'Activar'
      on Press: SetTag("DB_OP.RC1", 30); SetBit("DB_OP.OP_SELMANU1")
      Visibility <- "MANU"
      Appearance <- "DB_OP.RC1"
   Button "Botón_25" at 1145,523 size 72x33; TextOff 'Desactivar'
      on Press: SetTag("DB_OP.RC1", 31); SetBit("DB_OP.OP_SELMANU1")
      Visibility <- "MANU"
      Appearance <- "DB_OP.RC1"
   Button "Botón_14" at 1065,569 size 72x33; TextOff 'Activar'
      on Press: SetTag("DB_OP.RC1", 22); SetBit("DB_OP.OP_SELMANU1")
      Visibility <- "MANU"
      Appearance <- "DB_OP.RC1"
   Button "Botón_15" at 1065,606 size 72x33; TextOff 'Activar'
      on Press: SetTag("DB_OP.RC1", 24); SetBit("DB_OP.OP_SELMANU1")
      Visibility <- "MANU"
      Appearance <- "DB_OP.RC1"
   Button "Botón_16" at 1065,644 size 72x33; TextOff 'Activar'
      on Press: SetTag("DB_OP.RC1", 26); SetBit("DB_OP.OP_SELMANU1")
      Visibility <- "MANU"
      Appearance <- "DB_OP.RC1"
   Button "Botón_18" at 1145,569 size 72x33; TextOff 'Desactivar'
      on Press: SetTag("DB_OP.RC1", 23); SetBit("DB_OP.OP_SELMANU1")
      Visibility <- "MANU"
      Appearance <- "DB_OP.RC1"
   Button "Botón_19" at 1145,606 size 72x33; TextOff 'Desactivar'
      on Press: SetTag("DB_OP.RC1", 25); SetBit("DB_OP.OP_SELMANU1")
      Visibility <- "MANU"
      Appearance <- "DB_OP.RC1"
   Button "Botón_20" at 1145,644 size 72x33; TextOff 'Desactivar'
      on Press: SetTag("DB_OP.RC1", 27); SetBit("DB_OP.OP_SELMANU1")
      Visibility <- "MANU"
      Appearance <- "DB_OP.RC1"
   Rectangle "Rectángulo_10" at 988,26 size 248x201
      Visibility <- "MANU"
   Button "Botón_6" at 1012,65 size 202x33; TextOff 'Subir (Pistón Superior)'
      on Press: SetTag("DB_OP.RC1", 16); SetBit("DB_OP.OP_SELMANU1")
      Visibility <- "MANU"
      Appearance <- "DB_OP.RC1"
   Button "Botón_7" at 1012,103 size 202x33; TextOff 'Bajar (Pistón Superior)'
      on Press: SetTag("DB_OP.RC1", 15); SetBit("DB_OP.OP_SELMANU1")
      Visibility <- "MANU"
      Appearance <- "DB_OP.RC1"
   Button "Botón_8" at 1012,179 size 202x33; TextOff 'Bajar (Pistón Inferior)'
      on Press: SetTag("DB_OP.RC1", 13); SetBit("DB_OP.OP_SELMANU1")
      Visibility <- "MANU"
      Appearance <- "DB_OP.RC1"
   Button "Botón_9" at 1012,141 size 202x33; TextOff 'Subir (Pistón Inferior)'
      on Press: SetTag("DB_OP.RC1", 14); SetBit("DB_OP.OP_SELMANU1")
      Visibility <- "MANU"
      Appearance <- "DB_OP.RC1"
   Rectangle "Rectángulo_11" at 988,26 size 248x29
      Visibility <- "MANU"
   TextField "Campo de texto_7" at 1056,30 size 110x18; Text 'Movimiento Vertical'
      Visibility <- "MANU"
   GraphicIOField "Campo ES gráfico_1" at 159,226 size 460x334; PictureList "Araña"
      ProcessValue <- "Alarma_Araña"

PopupScreen "Comandos Almacenes" 1280x714
   Rectangle "Rectángulo_9" at 844,194 size 118x128
      Visibility <- "MANU"
   Rectangle "Rectángulo_8" at 844,194 size 118x29
      Visibility <- "MANU"
   TextField "Campo de texto_3" at 860,198 size 86x18; Text 'Intercambiador'
      Visibility <- "MANU"
   Button "Botón_1" at 859,238 size 88x33; TextOff 'Avance'
      on Press: SetTag("DB_OP.RC1", 1); SetBit("DB_OP.OP_SELMANU1")
      Visibility <- "MANU"
      Appearance <- "DB_OP.RC1"
   Button "Botón_2" at 859,276 size 88x33; TextOff 'Retroceso'
      on Press: SetTag("DB_OP.RC1", 2); SetBit("DB_OP.OP_SELMANU1")
      Visibility <- "MANU"
      Appearance <- "DB_OP.RC1"
   Circle "Cercle_1" at 407,425 size 14x14
      Appearance <- "26S6"
   TextField "Campo de texto_2" at 87,557 size 259x22; Text '26S7 - Almacén 2 en puesto de Espera'
   TextField "Campo de texto_4" at 36,478 size 266x22; Text '26S6 - Almacén 2 en puesto de Trabajo'
   GraphicIOField "Campo ES gráfico_2" at 416,233 size 388x286; PictureList "Grupo 1 - Almacén A"
      ProcessValue <- "26S7"
   GraphicIOField "Campo ES gráfico_1" at 416,233 size 388x286; PictureList "Grupo 1 - Almacén B"
      ProcessValue <- "26S7"
      Visibility <- "Alarma_Almacenes"
   Circle "Cercle_2" at 502,466 size 14x14
      Appearance <- "26S7"
   TextField "Campo de texto_6" at 52,590 size 285x22; Text 'M01 - Motor Intercambiador de Almacenes'

PopupScreen "Comandos Rolos" 1280x714
   GraphicIOField "Campo ES gráfico_4" at 134,166 size 538x272; PictureList "Rolos"
      ProcessValue <- "Alarma_Perfiladores"
   Polygon "Polígono_3" at 184,215 size 385x136
      Visibility <- "Rolos\Rolos.PresenciaPieza"
   Rectangle "Rectángulo_9" at 811,197 size 118x128
      Visibility <- "MANU"
   Rectangle "Rectángulo_8" at 811,197 size 118x29
      Visibility <- "MANU"
   TextField "Campo de texto_3" at 854,201 size 32x18; Text 'Rolos'
      Visibility <- "MANU"
   Button "Botón_29" at 826,241 size 88x33; TextOff 'Avance'
      on Press: SetTag("DB_OP.RC1", 41); SetBit("DB_OP.OP_SELMANU1")
      Visibility <- "MANU"
      Appearance <- "DB_OP.RC1"
   Button "Botón_30" at 826,279 size 88x33; TextOff 'Retroceso'
      on Press: SetTag("DB_OP.RC1", 42); SetBit("DB_OP.OP_SELMANU1")
      Visibility <- "MANU"
      Appearance <- "DB_OP.RC1"
   TextField "Campo de texto_7" at 303,476 size 104x32; Text '27S3 - Chapa en Entrada Perfilador'
   Circle "Cercle_10" at 201,328 size 12x12
      Appearance <- "27S3"
   Circle "Cercle_13" at 349,283 size 12x12
      Appearance <- "26S8"
   TextField "Campo de texto_11" at 455,437 size 114x32; Text '26S8 - Chapa en Transporte de Rolos'

PopupScreen "Comandos Piqueteador" 1280x714
   Button "Botón_32" at 397,449 size 118x33; TextOff 'Bajar Tope'
      on Press: SetTag("DB_OP.RC2", 36); SetBit("DB_OP.OP_SELMANU2")
      Visibility <- "MANU"
      Appearance <- "DB_OP.RC2"
   Button "Botón_33" at 397,411 size 118x33; TextOff 'Subir Tope'
      on Press: SetTag("DB_OP.RC2", 35); SetBit("DB_OP.OP_SELMANU2")
      Visibility <- "MANU"
      Appearance <- "DB_OP.RC2"
   Button "Botón_34" at 517,449 size 104x33; TextOff 'Bajar Herr.'
      on Press: SetTag("DB_OP.RC2", 40); SetBit("DB_OP.OP_SELMANU2")
      Visibility <- "MANU"
      Appearance <- "DB_OP.RC2"
   Button "Botón_35" at 517,411 size 104x33; TextOff 'Subir Herr.'
      on Press: SetTag("DB_OP.RC2", 41); SetBit("DB_OP.OP_SELMANU2")
      Visibility <- "MANU"
      Appearance <- "DB_OP.RC2"
   TextField "Campo de texto_5" at 1020,369 size 81x18; Text 'Herramienta 2'
   TextField "Campo de texto_2" at 748,373 size 81x18; Text 'Herramienta 1'
   Button "Botón_20" at 674,411 size 88x33; TextOff 'ON'
      on Press: SetTag("DB_OP.RC2", 42); SetBit("DB_OP.OP_SELMANU2")
      Visibility <- "MANU"
      Appearance <- "DB_OP.RC2"
   Button "Botón_21" at 946,411 size 88x33; TextOff 'ON'
      on Press: SetTag("DB_OP.RC2", 46); SetBit("DB_OP.OP_SELMANU2")
      Visibility <- "MANU"
      Appearance <- "DB_OP.RC2"
   Button "Botón_22" at 764,411 size 88x33; TextOff 'OFF'
      on Press: SetTag("DB_OP.RC2", 43); SetBit("DB_OP.OP_SELMANU2")
      Visibility <- "MANU"
      Appearance <- "DB_OP.RC2"
   Button "Botón_23" at 1036,411 size 88x33; TextOff 'OFF'
      on Press: SetTag("DB_OP.RC2", 47); SetBit("DB_OP.OP_SELMANU2")
      Visibility <- "MANU"
      Appearance <- "DB_OP.RC2"
   Button "Botón_28" at 674,449 size 88x33; TextOff 'ON'
      on Press: SetTag("DB_OP.RC2", 44); SetBit("DB_OP.OP_SELMANU2")
      Visibility <- "MANU"
      Appearance <- "DB_OP.RC2"
   Button "Botón_1" at 946,447 size 88x33; TextOff 'ON'
      on Press: SetTag("DB_OP.RC2", 48); SetBit("DB_OP.OP_SELMANU2")
      Visibility <- "MANU"
      Appearance <- "DB_OP.RC2"
   Button "Botón_2" at 764,449 size 88x33; TextOff 'OFF'
      on Press: SetTag("DB_OP.RC2", 45); SetBit("DB_OP.OP_SELMANU2")
      Visibility <- "MANU"
      Appearance <- "DB_OP.RC2"
   Button "Botón_31" at 1036,447 size 88x33; TextOff 'OFF'
      on Press: SetTag("DB_OP.RC2", 49); SetBit("DB_OP.OP_SELMANU2")
      Visibility <- "MANU"
      Appearance <- "DB_OP.RC2"
   GraphicIOField "Campo ES gráfico_8" at 250,43 size 289x268; PictureList "Formador"
      ProcessValue <- "Alarma_Formador"
   Rectangle "Rectángulo_9" at 930,366 size 254x128
      Visibility <- "MANU"
   Circle "Cercle_6" at 349,49 size 10x10
      Appearance <- "28S5"
   Circle "Cercle_7" at 349,78 size 10x10
      Appearance <- "28S6"
   TextField "Campo de texto_4" at 72,33 size 180x18; Text '28S5 - Herramientas Bloqueadas'
   TextField "Campo de texto_9" at 54,61 size 200x18; Text '28S6 - Herramientas Desbloqueadas'
   Circle "Cercle_8" at 451,121 size 10x10
      Appearance <- "28S3"
   Circle "Cercle_9" at 465,130 size 10x10
      Appearance <- "28S4"
   Circle "Cercle_10" at 518,168 size 10x10
      Appearance <- "28S1"
   Circle "Cercle_16" at 495,149 size 10x10
      Appearance <- "28S2"
   Circle "Cercle_0" at 433,216 size 10x10
      Appearance <- "27S5"
   Circle "Cercle_17" at 410,198 size 10x10
      Appearance <- "27S6"
   Circle "Cercle_18" at 361,163 size 10x10
      Appearance <- "27S7"
   Circle "Cercle_19" at 379,176 size 10x10
      Appearance <- "27S8"
   TextField "Campo de texto_14" at 530,72 size 146x18; Text '28S3 - Herr. 2 Matriz OFF'
   TextField "Campo de texto_15" at 543,91 size 142x18; Text '28S4 - Herr. 2 Matriz ON'
   TextField "Campo de texto_16" at 589,139 size 152x18; Text '28S1 - Herr. 2 Martillo OFF'
   TextField "Campo de texto_17" at 562,118 size 148x18; Text '28S2 - Herr. 2 Martillo ON'
   TextField "Campo de texto_18" at 40,196 size 146x18; Text '27S7 - Herr. 1 Matriz OFF'
   TextField "Campo de texto_19" at 64,219 size 142x18; Text '27S8 - Herr. 1 Matriz ON'
   TextField "Campo de texto_20" at 90,276 size 152x18; Text '27S5 - Herr. 1 Martillo OFF'
   TextField "Campo de texto_21" at 73,257 size 148x18; Text '27S6 - Herr. 1 Martillo ON'
   Rectangle "Rectángulo_1" at 381,369 size 254x128
      Visibility <- "MANU"
   Rectangle "Rectángulo_2" at 381,369 size 254x29
      Visibility <- "MANU"
   TextField "Campo de texto_1" at 491,373 size 45x18; Text 'General'
      Visibility <- "MANU"
   Rectangle "Rectángulo_3" at 658,369 size 254x128
      Visibility <- "MANU"
   IOField "Campo ES_1" at 480,552 size 96x32; FormatPattern 99999999
      ProcessValue <- "PosiciónFormado1"
   IOField "Campo ES_2" at 707,585 size 96x32; FormatPattern 99999999
      ProcessValue <- "PosiciónFormado2"
   IOField "Campo ES_3" at 480,585 size 96x32; FormatPattern 99999999
      ProcessValue <- "PosiciónFormado3"
   IOField "Campo ES_4" at 707,552 size 96x32; FormatPattern 99999999
      ProcessValue <- "PosiciónFormado4"
   TextField "Campo de texto_8" at 233,557 size 155x18; Text 'Posición para Herramienta 1'
   GraphicView "Visor de gráficos_1" at 701,252 size 114x83; Picture "a_4"
   GraphicView "Visor de gráficos_2" at 972,251 size 114x83; Picture "b_2"
   GraphicView "Visor de gráficos_3" at 1022,197 size 114x83; Picture "c_1"
   GraphicView "Visor de gráficos_4" at 751,198 size 114x83; Picture "b_2"
   TextField "Campo de texto_22" at 857,426 size 41x18; Text 'Martillo'
      Visibility <- "MANU"
   TextField "Campo de texto_23" at 857,455 size 35x18; Text 'Matriz'
      Visibility <- "MANU"
   TextField "Campo de texto_24" at 1129,426 size 41x18; Text 'Martillo'
      Visibility <- "MANU"
   TextField "Campo de texto_25" at 1129,455 size 35x18; Text 'Matriz'
      Visibility <- "MANU"
   TextField "Campo de texto_3" at 504,662 size 51x18; Text 'Corner 1'
   TextField "Campo de texto_6" at 233,589 size 155x18; Text 'Posición para Herramienta 2'
   TextField "Campo de texto_7" at 812,557 size 155x18; Text 'Posición para Herramienta 1'
   TextField "Campo de texto_10" at 812,589 size 155x18; Text 'Posición para Herramienta 2'
   TextField "Campo de texto_11" at 731,661 size 51x18; Text 'Corner 2'
   TextField "Campo de texto_12" at 394,557 size 80x18; Text 'Ajuste con F1'
   TextField "Campo de texto_13" at 394,589 size 80x18; Text 'Ajuste con F2'
   TextField "Campo de texto_26" at 970,557 size 80x18; Text 'Ajuste con F3'
   TextField "Campo de texto_27" at 970,589 size 80x18; Text 'Ajuste con F4'

